   "Carrier_33_Status.10" AT %I2001.2 : Bool;
   "Carrier_33_Status.11" AT %I2001.3 : Bool;
   "Carrier_33_Status.12" AT %I2001.4 : Bool;
   "Carrier_33_Status.13" AT %I2001.5 : Bool;
   "Carrier_33_Status.14" AT %I2001.6 : Bool;
   "Carrier_33_Status.15" AT %I2001.7 : Bool;
   "Carrier_33_SDCFaultCode" AT %IW2002 : Word;   // SDC FAULT CODE
   "Carrier_33_CarrierPosition" AT %ID2004 : DWord;   // CARRIER POSITION
   "Carrier_33_CarrierNumber" AT %IW2008 : Word;   // CARRIER NUMBER
   "Carrier_33_G120DControlWord" AT %IW2010 : Word;   // G120D_STW1_CONTROL
   "Carrier_33_G120DControlWord.0" AT %I2010.0 : Bool;   // Bit_00_ON
   "Carrier_33_G120DControlWord.1" AT %I2010.1 : Bool;   // Bit_01_AUS2_INH
   "Carrier_33_G120DControlWord.2" AT %I2010.2 : Bool;   // Bit_02_AUS3_STOP
   "Carrier_33_G120DControlWord.3" AT %I2010.3 : Bool;   // Bit_03_EN
   "Carrier_33_G120DControlWord.4" AT %I2010.4 : Bool;   // Bit_04_EN_RAMP
   "Carrier_33_G120DControlWord.5" AT %I2010.5 : Bool;   // Bit_05_START_RAMP
   "Carrier_33_G120DControlWord.6" AT %I2010.6 : Bool;   // Bit_06_SETPOINT
   "Carrier_33_G120DControlWord.7" AT %I2010.7 : Bool;   // Bit_07_RESET
   "Carrier_33_G120DControlWord.8" AT %I2011.0 : Bool;   // Bit_08_JOG_R
   "Carrier_33_G120DControlWord.9" AT %I2011.1 : Bool;   // Bit_09_JOG_L
   "Carrier_33_G120DControlWord.10" AT %I2011.2 : Bool;   // Bit_10_CONTR_PLC
   "Carrier_33_G120DControlWord.11" AT %I2011.3 : Bool;   // Bit_11_REVERSE
   "Carrier_33_G120DControlWord.12" AT %I2011.4 : Bool;   // Bit_12_BRAKE_RELEASE
   "Carrier_33_G120DControlWord.13" AT %I2011.5 : Bool;   // Bit_13_DDS
   "Carrier_33_G120DControlWord.14" AT %I2011.6 : Bool;   // Bit_14_DO0
   "Carrier_33_G120DControlWord.15" AT %I2011.7 : Bool;   // Bit_15_DO1
   "Carrier_33_G120DStatusWord" AT %IW2012 : Word;   // G120D_ZSW1_STATUS
   "Carrier_33_G120DStatusWord.0" AT %I2012.0 : Bool;   // Bit_00_READY_RUN
   "Carrier_33_G120DStatusWord.1" AT %I2012.1 : Bool;   // Bit_01_READY_ON
   "Carrier_33_G120DStatusWord.2" AT %I2012.2 : Bool;   // Bit_02_ENABLE
   "Carrier_33_G120DStatusWord.3" AT %I2012.3 : Bool;   // Bit_03_FAULT
   "Carrier_33_G120DStatusWord.4" AT %I2012.4 : Bool;   // Bit_04_OFF2
   "Carrier_33_G120DStatusWord.5" AT %I2012.5 : Bool;   // Bit_05_OFF3
   "Carrier_33_G120DStatusWord.6" AT %I2012.6 : Bool;   // Bit_06_LOCK_OUT
   "Carrier_33_G120DStatusWord.7" AT %I2012.7 : Bool;   // Bit_07_WARN
   "Carrier_33_G120DStatusWord.8" AT %I2013.0 : Bool;   // Bit_08_NO_DEVIATION
   "Carrier_33_G120DStatusWord.9" AT %I2013.1 : Bool;   // Bit_09_CONTR_PLC
   "Carrier_33_G120DStatusWord.10" AT %I2013.2 : Bool;   // Bit_10_F_MAX
   "Carrier_33_G120DStatusWord.11" AT %I2013.3 : Bool;   // Bit_11_LIMIT_REACHED
   "Carrier_33_G120DStatusWord.12" AT %I2013.4 : Bool;   // Bit_12_BRAKE_OPEN
   "Carrier_33_G120DStatusWord.13" AT %I2013.5 : Bool;   // Bit_13_NO_OVERTEMP
   "Carrier_33_G120DStatusWord.14" AT %I2013.6 : Bool;   // Bit_14_CW_CCW
   "Carrier_33_G120DStatusWord.15" AT %I2013.7 : Bool;   // Bit_15_OVERL
   "Carrier_33_Slot2_Input" AT %IW2014 : Word;   // SLOT 2 INPUT WORD
   "Carrier_33_CrashDetectSW" AT %I2014.0 : Bool;   // CRASH DETECT SW
   "Carrier_33_SpareSafetyInput(2_1)" AT %I2014.1 : Bool;   // SPARE SAFETY INPUT
   "Carrier_33_SpareSafetyInput(2_2)" AT %I2014.2 : Bool;   // SPARE SAFETY INPUT
   "Carrier_33_SpareSafetyInput(2_3)" AT %I2014.3 : Bool;   // SPARE SAFETY INPUT
   "Carrier_33_SpareSafetyInput(2_4)" AT %I2014.4 : Bool;   // SPARE SAFETY INPUT
   "Carrier_33_SpareSafetyInput(2_5)" AT %I2014.5 : Bool;   // SPARE SAFETY INPUT
   "Carrier_33_SpareSafetyInput(2_6)" AT %I2014.6 : Bool;   // SPARE SAFETY INPUT
   "Carrier_33_SpareSafetyInput(2_7)" AT %I2014.7 : Bool;   // SPARE SAFETY INPUT
   "Carrier_33_Slot3_SafetyOutput" AT %IW2015 : Word;   // SLOT 3 SAFETY OUTPUT WORD
   "Carrier_33_Crash_Detect_OK" AT %I2015.0 : Bool;   // CARRIER CRASH DETECT
   "Carrier_33_SpareSafetyOutput(3_1)" AT %I2015.1 : Bool;   // SPARE SAFETY OUTPUT
   "Carrier_33_SpareSafetyOutput(3_2)" AT %I2015.2 : Bool;   // SPARE SAFETY OUTPUT
   "Carrier_33_SpareSafetyOutput(3_3)" AT %I2015.3 : Bool;   // SPARE SAFETY OUTPUT
   "Carrier_33_SpareSafetyOutput(3_4)" AT %I2015.4 : Bool;   // SPARE SAFETY OUTPUT
   "Carrier_33_SpareSafetyOutput(3_5)" AT %I2015.5 : Bool;   // SPARE SAFETY OUTPUT
   "Carrier_33_SpareSafetyOutput(3_6)" AT %I2015.6 : Bool;   // SPARE SAFETY OUTPUT
   "Carrier_33_SpareSafetyOutput(3_7)" AT %I2015.7 : Bool;   // SPARE SAFETY OUTPUT
   "Carrier_33_Slot4_Input" AT %IW2016 : Word;   // SLOT 4 INPUT WORD
   "Carrier_33_480VPowerOn_MDCB1" AT %I2016.0 : Bool;   // 480 VAC POWER ON MDCB 1
   "Carrier_33_SpareInput(4_1)" AT %I2016.1 : Bool;   // SPARE INPUT
   "Carrier_33_SpareInput(4_2)" AT %I2016.2 : Bool;   // SPARE INPUT
   "Carrier_33_SitopSelectStatus" AT %I2016.3 : Bool;   // SITOP SELECT STATUS
   "Carrier_33_DCsupplyOnPSCB2" AT %I2016.4 : Bool;   // DC SUPPLY ON PSCB 2
   "Carrier_33_SpareInput(4_5)" AT %I2016.5 : Bool;   // SPARE INPUT
   "Carrier_33_SpareInput(4_6)" AT %I2016.6 : Bool;   // SPARE INPUT
   "Carrier_33_SpareInput(4_7)" AT %I2016.7 : Bool;   // SPARE INPUT
   "Carrier_33_PB1_ProdHoldLH" AT %I2017.0 : Bool;   // PB 1 PRODUCTION HOLD LH
   "Carrier_33_PB2_ResetLH" AT %I2017.1 : Bool;   // PB 2 RESET LH
   "Carrier_33_PB3_ProdHoldRH" AT %I2017.2 : Bool;   // PB 3 PRODUCTION HOLD RH
   "Carrier_33_PB4_ResetRH" AT %I2017.3 : Bool;   // PB 4 RESET RH
   "Carrier_33_SpareInput(4_14)" AT %I2017.4 : Bool;   // SPARE INPUT
   "Carrier_33_SpareInput(4_15)" AT %I2017.5 : Bool;   // SPARE INPUT
   "Carrier_33_SpareInput(4_16)" AT %I2017.6 : Bool;   // SPARE INPUT
   "Carrier_33_SpareInput(4_17)" AT %I2017.7 : Bool;   // SPARE INPUT
   "Carrier_33_Slot5_Output" AT %IW2018 : Word;   // SLOT 5 OUTPUT WORD
   "Carrier_33_IRD400_HMI_24VDC_ENABLE" AT %I2018.0 : Bool;   // IRD 400 PANEL HMI 24V DC POWER
   "Carrier_33_FaultLight_LH" AT %I2018.1 : Bool;   // FAULT LIGHT LH
   "Carrier_33_RunLight_LH" AT %I2018.2 : Bool;   // RUN LIGHT LH
   "Carrier_33_FaultLight_RH" AT %I2018.3 : Bool;   // FAULT LIGHT RH
   "Carrier_33_RunLight_RH" AT %I2018.4 : Bool;   // RUN LIGHT RH
   "Carrier_33_SpareOutput(5_5)" AT %I2018.5 : Bool;   // SPARE OUTPUT
   "Carrier_33_SpareOutput(5_6)" AT %I2018.6 : Bool;   // SPARE OUTPUT
   "Carrier_33_SpareOutput(5_7)" AT %I2018.7 : Bool;   // SPARE OUTPUT
   "Carrier_33_ActualSpeed" AT %IW2020 : Word;   // ACTUAL SPEED
   "Carrier_33_CarrierDriveAlarm" AT %IW2022 : Word;   // CARRIER DRIVE ALARM
   "Carrier_33_CarrierDriveWarning" AT %IW2024 : Word;   // CARRIER DRIVE WARNING
   "Carrier_34_Status" AT %IW2050 : Word;   // CARRIER STATUS WORD
   "Carrier_34_Status.0" AT %I2050.0 : Bool;   // HEARTBEAT
   "Carrier_34_Status.1" AT %I2050.1 : Bool;   // MANUAL
   "Carrier_34_Status.2" AT %I2050.2 : Bool;   // IN_AUTO
   "Carrier_34_Status.3" AT %I2050.3 : Bool;   // POSITIONING_COMPLETE
   "Carrier_34_Status.4" AT %I2050.4 : Bool;   // PRODUCTION HOLD
   "Carrier_34_Status.5" AT %I2050.5 : Bool;   // CARRIER MOVING FORWARD
   "Carrier_34_Status.6" AT %I2050.6 : Bool;   // CARRIER MOVING REVERSE
   "Carrier_34_Status.7" AT %I2050.7 : Bool;   // CARRIER FAULT
   "Carrier_34_Status.8" AT %I2051.0 : Bool;   // CRASH DETECT TRIPPED
   "Carrier_34_Status.9" AT %I2051.1 : Bool;
   "Carrier_34_Status.10" AT %I2051.2 : Bool;
   "Carrier_34_Status.11" AT %I2051.3 : Bool;
   "Carrier_34_Status.12" AT %I2051.4 : Bool;
   "Carrier_34_Status.13" AT %I2051.5 : Bool;
   "Carrier_34_Status.14" AT %I2051.6 : Bool;
   "Carrier_34_Status.15" AT %I2051.7 : Bool;
   "Carrier_34_SDCFaultCode" AT %IW2052 : Word;   // SDC FAULT CODE
   "Carrier_34_CarrierPosition" AT %ID2054 : DWord;   // CARRIER POSITION
   "Carrier_34_CarrierNumber" AT %IW2058 : Word;   // CARRIER NUMBER
   "Carrier_34_G120DControlWord" AT %IW2060 : Word;   // G120D_STW1_CONTROL
   "Carrier_34_G120DControlWord.0" AT %I2060.0 : Bool;   // Bit_00_ON
   "Carrier_34_G120DControlWord.1" AT %I2060.1 : Bool;   // Bit_01_AUS2_INH
   "Carrier_34_G120DControlWord.2" AT %I2060.2 : Bool;   // Bit_02_AUS3_STOP
   "Carrier_34_G120DControlWord.3" AT %I2060.3 : Bool;   // Bit_03_EN
   "Carrier_34_G120DControlWord.4" AT %I2060.4 : Bool;   // Bit_04_EN_RAMP
   "Carrier_34_G120DControlWord.5" AT %I2060.5 : Bool;   // Bit_05_START_RAMP
   "Carrier_34_G120DControlWord.6" AT %I2060.6 : Bool;   // Bit_06_SETPOINT
   "Carrier_34_G120DControlWord.7" AT %I2060.7 : Bool;   // Bit_07_RESET
   "Carrier_34_G120DControlWord.8" AT %I2061.0 : Bool;   // Bit_08_JOG_R
   "Carrier_34_G120DControlWord.9" AT %I2061.1 : Bool;   // Bit_09_JOG_L
   "Carrier_34_G120DControlWord.10" AT %I2061.2 : Bool;   // Bit_10_CONTR_PLC
   "Carrier_34_G120DControlWord.11" AT %I2061.3 : Bool;   // Bit_11_REVERSE
   "Carrier_34_G120DControlWord.12" AT %I2061.4 : Bool;   // Bit_12_BRAKE_RELEASE
   "Carrier_34_G120DControlWord.13" AT %I2061.5 : Bool;   // Bit_13_DDS
   "Carrier_34_G120DControlWord.14" AT %I2061.6 : Bool;   // Bit_14_DO0
   "Carrier_34_G120DControlWord.15" AT %I2061.7 : Bool;   // Bit_15_DO1
   "Carrier_34_G120DStatusWord" AT %IW2062 : Word;   // G120D_ZSW1_STATUS
   "Carrier_34_G120DStatusWord.0" AT %I2062.0 : Bool;   // Bit_00_READY_RUN
   "Carrier_34_G120DStatusWord.1" AT %I2062.1 : Bool;   // Bit_01_READY_ON
   "Carrier_34_G120DStatusWord.2" AT %I2062.2 : Bool;   // Bit_02_ENABLE
   "Carrier_34_G120DStatusWord.3" AT %I2062.3 : Bool;   // Bit_03_FAULT
   "Carrier_34_G120DStatusWord.4" AT %I2062.4 : Bool;   // Bit_04_OFF2
   "Carrier_34_G120DStatusWord.5" AT %I2062.5 : Bool;   // Bit_05_OFF3
   "Carrier_34_G120DStatusWord.6" AT %I2062.6 : Bool;   // Bit_06_LOCK_OUT
   "Carrier_34_G120DStatusWord.7" AT %I2062.7 : Bool;   // Bit_07_WARN
   "Carrier_34_G120DStatusWord.8" AT %I2063.0 : Bool;   // Bit_08_NO_DEVIATION
   "Carrier_34_G120DStatusWord.9" AT %I2063.1 : Bool;   // Bit_09_CONTR_PLC
   "Carrier_34_G120DStatusWord.10" AT %I2063.2 : Bool;   // Bit_10_F_MAX
   "Carrier_34_G120DStatusWord.11" AT %I2063.3 : Bool;   // Bit_11_LIMIT_REACHED
   "Carrier_34_G120DStatusWord.12" AT %I2063.4 : Bool;   // Bit_12_BRAKE_OPEN
   "Carrier_34_G120DStatusWord.13" AT %I2063.5 : Bool;   // Bit_13_NO_OVERTEMP
   "Carrier_34_G120DStatusWord.14" AT %I2063.6 : Bool;   // Bit_14_CW_CCW
   "Carrier_34_G120DStatusWord.15" AT %I2063.7 : Bool;   // Bit_15_OVERL
   "Carrier_34_Slot2_Input" AT %IW2064 : Word;   // SLOT 2 INPUT WORD
   "Carrier_34_CrashDetectSW" AT %I2064.0 : Bool;   // CRASH DETECT SW
   "Carrier_34_SpareSafetyInput(2_1)" AT %I2064.1 : Bool;   // SPARE SAFETY INPUT
   "Carrier_34_SpareSafetyInput(2_2)" AT %I2064.2 : Bool;   // SPARE SAFETY INPUT
   "Carrier_34_SpareSafetyInput(2_3)" AT %I2064.3 : Bool;   // SPARE SAFETY INPUT
   "Carrier_34_SpareSafetyInput(2_4)" AT %I2064.4 : Bool;   // SPARE SAFETY INPUT
   "Carrier_34_SpareSafetyInput(2_5)" AT %I2064.5 : Bool;   // SPARE SAFETY INPUT
   "Carrier_34_SpareSafetyInput(2_6)" AT %I2064.6 : Bool;   // SPARE SAFETY INPUT
   "Carrier_34_SpareSafetyInput(2_7)" AT %I2064.7 : Bool;   // SPARE SAFETY INPUT
   "Carrier_34_Slot3_SafetyOutput" AT %IW2065 : Word;   // SLOT 3 SAFETY OUTPUT WORD
   "Carrier_34_Crash_Detect_OK" AT %I2065.0 : Bool;   // CARRIER CRASH DETECT
   "Carrier_34_SpareSafetyOutput(3_1)" AT %I2065.1 : Bool;   // SPARE SAFETY OUTPUT
   "Carrier_34_SpareSafetyOutput(3_2)" AT %I2065.2 : Bool;   // SPARE SAFETY OUTPUT
   "Carrier_34_SpareSafetyOutput(3_3)" AT %I2065.3 : Bool;   // SPARE SAFETY OUTPUT
   "Carrier_34_SpareSafetyOutput(3_4)" AT %I2065.4 : Bool;   // SPARE SAFETY OUTPUT
   "Carrier_34_SpareSafetyOutput(3_5)" AT %I2065.5 : Bool;   // SPARE SAFETY OUTPUT
   "Carrier_34_SpareSafetyOutput(3_6)" AT %I2065.6 : Bool;   // SPARE SAFETY OUTPUT
   "Carrier_34_SpareSafetyOutput(3_7)" AT %I2065.7 : Bool;   // SPARE SAFETY OUTPUT
   "Carrier_34_Slot4_Input" AT %IW2066 : Word;   // SLOT 4 INPUT WORD
   "Carrier_34_480VPowerOn_MDCB1" AT %I2066.0 : Bool;   // 480 VAC POWER ON MDCB 1
   "Carrier_34_SpareInput(4_1)" AT %I2066.1 : Bool;   // SPARE INPUT
   "Carrier_34_SpareInput(4_2)" AT %I2066.2 : Bool;   // SPARE INPUT
   "Carrier_34_SitopSelectStatus" AT %I2066.3 : Bool;   // SITOP SELECT STATUS
   "Carrier_34_DCsupplyOnPSCB2" AT %I2066.4 : Bool;   // DC SUPPLY ON PSCB 2
   "Carrier_34_SpareInput(4_5)" AT %I2066.5 : Bool;   // SPARE INPUT
   "Carrier_34_SpareInput(4_6)" AT %I2066.6 : Bool;   // SPARE INPUT
   "Carrier_34_SpareInput(4_7)" AT %I2066.7 : Bool;   // SPARE INPUT
   "Carrier_34_PB1_ProdHoldLH" AT %I2067.0 : Bool;   // PB 1 PRODUCTION HOLD LH
   "Carrier_34_PB2_ResetLH" AT %I2067.1 : Bool;   // PB 2 RESET LH
   "Carrier_34_PB3_ProdHoldRH" AT %I2067.2 : Bool;   // PB 3 PRODUCTION HOLD RH
   "Carrier_34_PB4_ResetRH" AT %I2067.3 : Bool;   // PB 4 RESET RH
   "Carrier_34_SpareInput(4_14)" AT %I2067.4 : Bool;   // SPARE INPUT
   "Carrier_34_SpareInput(4_15)" AT %I2067.5 : Bool;   // SPARE INPUT
   "Carrier_34_SpareInput(4_16)" AT %I2067.6 : Bool;   // SPARE INPUT
   "Carrier_34_SpareInput(4_17)" AT %I2067.7 : Bool;   // SPARE INPUT
   "Carrier_34_Slot5_Output" AT %IW2068 : Word;   // SLOT 5 OUTPUT WORD
   "Carrier_34_IRD400_HMI_24VDC_ENABLE" AT %I2068.0 : Bool;   // IRD 400 PANEL HMI 24V DC POWER
   "Carrier_34_FaultLight_LH" AT %I2068.1 : Bool;   // FAULT LIGHT LH
   "Carrier_34_RunLight_LH" AT %I2068.2 : Bool;   // RUN LIGHT LH
   "Carrier_34_FaultLight_RH" AT %I2068.3 : Bool;   // FAULT LIGHT RH
   "Carrier_34_RunLight_RH" AT %I2068.4 : Bool;   // RUN LIGHT RH
   "Carrier_34_SpareOutput(5_5)" AT %I2068.5 : Bool;   // SPARE OUTPUT
   "Carrier_34_SpareOutput(5_6)" AT %I2068.6 : Bool;   // SPARE OUTPUT
   "Carrier_34_SpareOutput(5_7)" AT %I2068.7 : Bool;   // SPARE OUTPUT
   "Carrier_34_ActualSpeed" AT %IW2070 : Word;   // ACTUAL SPEED
   "Carrier_34_CarrierDriveAlarm" AT %IW2072 : Word;   // CARRIER DRIVE ALARM
   "Carrier_34_CarrierDriveWarning" AT %IW2074 : Word;   // CARRIER DRIVE WARNING
   "Carrier_35_Status" AT %IW2100 : Word;   // CARRIER STATUS WORD
   "Carrier_35_Status.0" AT %I2100.0 : Bool;   // HEARTBEAT
   "Carrier_35_Status.1" AT %I2100.1 : Bool;   // MANUAL
   "Carrier_35_Status.2" AT %I2100.2 : Bool;   // IN_AUTO
   "Carrier_35_Status.3" AT %I2100.3 : Bool;   // POSITIONING_COMPLETE
   "Carrier_35_Status.4" AT %I2100.4 : Bool;   // PRODUCTION HOLD
   "Carrier_35_Status.5" AT %I2100.5 : Bool;   // CARRIER MOVING FORWARD
   "Carrier_35_Status.6" AT %I2100.6 : Bool;   // CARRIER MOVING REVERSE
   "Carrier_35_Status.7" AT %I2100.7 : Bool;   // CARRIER FAULT
   "Carrier_35_Status.8" AT %I2101.0 : Bool;   // CRASH DETECT TRIPPED
   "Carrier_35_Status.9" AT %I2101.1 : Bool;
   "Carrier_35_Status.10" AT %I2101.2 : Bool;
   "Carrier_35_Status.11" AT %I2101.3 : Bool;
   "Carrier_35_Status.12" AT %I2101.4 : Bool;
   "Carrier_35_Status.13" AT %I2101.5 : Bool;
   "Carrier_35_Status.14" AT %I2101.6 : Bool;
   "Carrier_35_Status.15" AT %I2101.7 : Bool;
   "Carrier_35_SDCFaultCode" AT %IW2102 : Word;   // SDC FAULT CODE
   "Carrier_35_CarrierPosition" AT %ID2104 : DWord;   // CARRIER POSITION
   "Carrier_35_CarrierNumber" AT %IW2108 : Word;   // CARRIER NUMBER
   "Carrier_35_G120DControlWord" AT %IW2110 : Word;   // G120D_STW1_CONTROL
   "Carrier_35_G120DControlWord.0" AT %I2110.0 : Bool;   // Bit_00_ON
   "Carrier_35_G120DControlWord.1" AT %I2110.1 : Bool;   // Bit_01_AUS2_INH
   "Carrier_35_G120DControlWord.2" AT %I2110.2 : Bool;   // Bit_02_AUS3_STOP
   "Carrier_35_G120DControlWord.3" AT %I2110.3 : Bool;   // Bit_03_EN
   "Carrier_35_G120DControlWord.4" AT %I2110.4 : Bool;   // Bit_04_EN_RAMP
   "Carrier_35_G120DControlWord.5" AT %I2110.5 : Bool;   // Bit_05_START_RAMP
   "Carrier_35_G120DControlWord.6" AT %I2110.6 : Bool;   // Bit_06_SETPOINT
   "Carrier_35_G120DControlWord.7" AT %I2110.7 : Bool;   // Bit_07_RESET
   "Carrier_35_G120DControlWord.8" AT %I2111.0 : Bool;   // Bit_08_JOG_R
   "Carrier_35_G120DControlWord.9" AT %I2111.1 : Bool;   // Bit_09_JOG_L
   "Carrier_35_G120DControlWord.10" AT %I2111.2 : Bool;   // Bit_10_CONTR_PLC
   "Carrier_35_G120DControlWord.11" AT %I2111.3 : Bool;   // Bit_11_REVERSE
   "Carrier_35_G120DControlWord.12" AT %I2111.4 : Bool;   // Bit_12_BRAKE_RELEASE
   "Carrier_35_G120DControlWord.13" AT %I2111.5 : Bool;   // Bit_13_DDS
   "Carrier_35_G120DControlWord.14" AT %I2111.6 : Bool;   // Bit_14_DO0
   "Carrier_35_G120DControlWord.15" AT %I2111.7 : Bool;   // Bit_15_DO1
   "Carrier_35_G120DStatusWord" AT %IW2112 : Word;   // G120D_ZSW1_STATUS
   "Carrier_35_G120DStatusWord.0" AT %I2112.0 : Bool;   // Bit_00_READY_RUN
   "Carrier_35_G120DStatusWord.1" AT %I2112.1 : Bool;   // Bit_01_READY_ON
   "Carrier_35_G120DStatusWord.2" AT %I2112.2 : Bool;   // Bit_02_ENABLE
   "Carrier_35_G120DStatusWord.3" AT %I2112.3 : Bool;   // Bit_03_FAULT
   "Carrier_35_G120DStatusWord.4" AT %I2112.4 : Bool;   // Bit_04_OFF2
   "Carrier_35_G120DStatusWord.5" AT %I2112.5 : Bool;   // Bit_05_OFF3
   "Carrier_35_G120DStatusWord.6" AT %I2112.6 : Bool;   // Bit_06_LOCK_OUT
   "Carrier_35_G120DStatusWord.7" AT %I2112.7 : Bool;   // Bit_07_WARN
   "Carrier_35_G120DStatusWord.8" AT %I2113.0 : Bool;   // Bit_08_NO_DEVIATION
   "Carrier_35_G120DStatusWord.9" AT %I2113.1 : Bool;   // Bit_09_CONTR_PLC
   "Carrier_35_G120DStatusWord.10" AT %I2113.2 : Bool;   // Bit_10_F_MAX
   "Carrier_35_G120DStatusWord.11" AT %I2113.3 : Bool;   // Bit_11_LIMIT_REACHED
   "Carrier_35_G120DStatusWord.12" AT %I2113.4 : Bool;   // Bit_12_BRAKE_OPEN
   "Carrier_35_G120DStatusWord.13" AT %I2113.5 : Bool;   // Bit_13_NO_OVERTEMP
   "Carrier_35_G120DStatusWord.14" AT %I2113.6 : Bool;   // Bit_14_CW_CCW
   "Carrier_35_G120DStatusWord.15" AT %I2113.7 : Bool;   // Bit_15_OVERL
   "Carrier_35_Slot2_Input" AT %IW2114 : Word;   // SLOT 2 INPUT WORD
   "Carrier_35_CrashDetectSW" AT %I2114.0 : Bool;   // CRASH DETECT SW
   "Carrier_35_SpareSafetyInput(2_1)" AT %I2114.1 : Bool;   // SPARE SAFETY INPUT
   "Carrier_35_SpareSafetyInput(2_2)" AT %I2114.2 : Bool;   // SPARE SAFETY INPUT
   "Carrier_35_SpareSafetyInput(2_3)" AT %I2114.3 : Bool;   // SPARE SAFETY INPUT
   "Carrier_35_SpareSafetyInput(2_4)" AT %I2114.4 : Bool;   // SPARE SAFETY INPUT
   "Carrier_35_SpareSafetyInput(2_5)" AT %I2114.5 : Bool;   // SPARE SAFETY INPUT
   "Carrier_35_SpareSafetyInput(2_6)" AT %I2114.6 : Bool;   // SPARE SAFETY INPUT
   "Carrier_35_SpareSafetyInput(2_7)" AT %I2114.7 : Bool;   // SPARE SAFETY INPUT
   "Carrier_35_Slot3_SafetyOutput" AT %IW2115 : Word;   // SLOT 3 SAFETY OUTPUT WORD
   "Carrier_35_Crash_Detect_OK" AT %I2115.0 : Bool;   // CARRIER CRASH DETECT
   "Carrier_35_SpareSafetyOutput(3_1)" AT %I2115.1 : Bool;   // SPARE SAFETY OUTPUT
   "Carrier_35_SpareSafetyOutput(3_2)" AT %I2115.2 : Bool;   // SPARE SAFETY OUTPUT
   "Carrier_35_SpareSafetyOutput(3_3)" AT %I2115.3 : Bool;   // SPARE SAFETY OUTPUT
   "Carrier_35_SpareSafetyOutput(3_4)" AT %I2115.4 : Bool;   // SPARE SAFETY OUTPUT
   "Carrier_35_SpareSafetyOutput(3_5)" AT %I2115.5 : Bool;   // SPARE SAFETY OUTPUT
   "Carrier_35_SpareSafetyOutput(3_6)" AT %I2115.6 : Bool;   // SPARE SAFETY OUTPUT
   "Carrier_35_SpareSafetyOutput(3_7)" AT %I2115.7 : Bool;   // SPARE SAFETY OUTPUT
   "Carrier_35_Slot4_Input" AT %IW2116 : Word;   // SLOT 4 INPUT WORD
   "Carrier_35_480VPowerOn_MDCB1" AT %I2116.0 : Bool;   // 480 VAC POWER ON MDCB 1
   "Carrier_35_SpareInput(4_1)" AT %I2116.1 : Bool;   // SPARE INPUT
   "Carrier_35_SpareInput(4_2)" AT %I2116.2 : Bool;   // SPARE INPUT
   "Carrier_35_SitopSelectStatus" AT %I2116.3 : Bool;   // SITOP SELECT STATUS
   "Carrier_35_DCsupplyOnPSCB2" AT %I2116.4 : Bool;   // DC SUPPLY ON PSCB 2
   "Carrier_35_SpareInput(4_5)" AT %I2116.5 : Bool;   // SPARE INPUT
   "Carrier_35_SpareInput(4_6)" AT %I2116.6 : Bool;   // SPARE INPUT
   "Carrier_35_SpareInput(4_7)" AT %I2116.7 : Bool;   // SPARE INPUT
   "Carrier_35_PB1_ProdHoldLH" AT %I2117.0 : Bool;   // PB 1 PRODUCTION HOLD LH
   "Carrier_35_PB2_ResetLH" AT %I2117.1 : Bool;   // PB 2 RESET LH
   "Carrier_35_PB3_ProdHoldRH" AT %I2117.2 : Bool;   // PB 3 PRODUCTION HOLD RH
   "Carrier_35_PB4_ResetRH" AT %I2117.3 : Bool;   // PB 4 RESET RH
   "Carrier_35_SpareInput(4_14)" AT %I2117.4 : Bool;   // SPARE INPUT
   "Carrier_35_SpareInput(4_15)" AT %I2117.5 : Bool;   // SPARE INPUT
   "Carrier_35_SpareInput(4_16)" AT %I2117.6 : Bool;   // SPARE INPUT
   "Carrier_35_SpareInput(4_17)" AT %I2117.7 : Bool;   // SPARE INPUT
   "Carrier_35_Slot5_Output" AT %IW2118 : Word;   // SLOT 5 OUTPUT WORD
   "Carrier_35_IRD400_HMI_24VDC_ENABLE" AT %I2118.0 : Bool;   // IRD 400 PANEL HMI 24V DC POWER
   "Carrier_35_FaultLight_LH" AT %I2118.1 : Bool;   // FAULT LIGHT LH
   "Carrier_35_RunLight_LH" AT %I2118.2 : Bool;   // RUN LIGHT LH
   "Carrier_35_FaultLight_RH" AT %I2118.3 : Bool;   // FAULT LIGHT RH
   "Carrier_35_RunLight_RH" AT %I2118.4 : Bool;   // RUN LIGHT RH
   "Carrier_35_SpareOutput(5_5)" AT %I2118.5 : Bool;   // SPARE OUTPUT
   "Carrier_35_SpareOutput(5_6)" AT %I2118.6 : Bool;   // SPARE OUTPUT
   "Carrier_35_SpareOutput(5_7)" AT %I2118.7 : Bool;   // SPARE OUTPUT
   "Carrier_35_ActualSpeed" AT %IW2120 : Word;   // ACTUAL SPEED
   "Carrier_35_CarrierDriveAlarm" AT %IW2122 : Word;   // CARRIER DRIVE ALARM
   "Carrier_35_CarrierDriveWarning" AT %IW2124 : Word;   // CARRIER DRIVE WARNING
   "Carrier_36_Status" AT %IW2150 : Word;   // CARRIER STATUS WORD
   "Carrier_36_Status.0" AT %I2150.0 : Bool;   // HEARTBEAT
   "Carrier_36_Status.1" AT %I2150.1 : Bool;   // MANUAL
   "Carrier_36_Status.2" AT %I2150.2 : Bool;   // IN_AUTO
   "Carrier_36_Status.3" AT %I2150.3 : Bool;   // POSITIONING_COMPLETE
   "Carrier_36_Status.4" AT %I2150.4 : Bool;   // PRODUCTION HOLD
   "Carrier_36_Status.5" AT %I2150.5 : Bool;   // CARRIER MOVING FORWARD
   "Carrier_36_Status.6" AT %I2150.6 : Bool;   // CARRIER MOVING REVERSE
   "Carrier_36_Status.7" AT %I2150.7 : Bool;   // CARRIER FAULT
   "Carrier_36_Status.8" AT %I2151.0 : Bool;   // CRASH DETECT TRIPPED
   "Carrier_36_Status.9" AT %I2151.1 : Bool;
   "Carrier_36_Status.10" AT %I2151.2 : Bool;
   "Carrier_36_Status.11" AT %I2151.3 : Bool;
   "Carrier_36_Status.12" AT %I2151.4 : Bool;
   "Carrier_36_Status.13" AT %I2151.5 : Bool;
   "Carrier_36_Status.14" AT %I2151.6 : Bool;
   "Carrier_36_Status.15" AT %I2151.7 : Bool;
   "Carrier_36_SDCFaultCode" AT %IW2152 : Word;   // SDC FAULT CODE
   "Carrier_36_CarrierPosition" AT %ID2154 : DWord;   // CARRIER POSITION
   "Carrier_36_CarrierNumber" AT %IW2158 : Word;   // CARRIER NUMBER
   "Carrier_36_G120DControlWord" AT %IW2160 : Word;   // G120D_STW1_CONTROL
   "Carrier_36_G120DControlWord.0" AT %I2160.0 : Bool;   // Bit_00_ON
   "Carrier_36_G120DControlWord.1" AT %I2160.1 : Bool;   // Bit_01_AUS2_INH
   "Carrier_36_G120DControlWord.2" AT %I2160.2 : Bool;   // Bit_02_AUS3_STOP
   "Carrier_36_G120DControlWord.3" AT %I2160.3 : Bool;   // Bit_03_EN
   "Carrier_36_G120DControlWord.4" AT %I2160.4 : Bool;   // Bit_04_EN_RAMP
   "Carrier_36_G120DControlWord.5" AT %I2160.5 : Bool;   // Bit_05_START_RAMP
   "Carrier_36_G120DControlWord.6" AT %I2160.6 : Bool;   // Bit_06_SETPOINT
   "Carrier_36_G120DControlWord.7" AT %I2160.7 : Bool;   // Bit_07_RESET
   "Carrier_36_G120DControlWord.8" AT %I2161.0 : Bool;   // Bit_08_JOG_R
   "Carrier_36_G120DControlWord.9" AT %I2161.1 : Bool;   // Bit_09_JOG_L
   "Carrier_36_G120DControlWord.10" AT %I2161.2 : Bool;   // Bit_10_CONTR_PLC
   "Carrier_36_G120DControlWord.11" AT %I2161.3 : Bool;   // Bit_11_REVERSE
   "Carrier_36_G120DControlWord.12" AT %I2161.4 : Bool;   // Bit_12_BRAKE_RELEASE
   "Carrier_36_G120DControlWord.13" AT %I2161.5 : Bool;   // Bit_13_DDS
   "Carrier_36_G120DControlWord.14" AT %I2161.6 : Bool;   // Bit_14_DO0
   "Carrier_36_G120DControlWord.15" AT %I2161.7 : Bool;   // Bit_15_DO1
   "Carrier_36_G120DStatusWord" AT %IW2162 : Word;   // G120D_ZSW1_STATUS
   "Carrier_36_G120DStatusWord.0" AT %I2162.0 : Bool;   // Bit_00_READY_RUN
   "Carrier_36_G120DStatusWord.1" AT %I2162.1 : Bool;   // Bit_01_READY_ON
   "Carrier_36_G120DStatusWord.2" AT %I2162.2 : Bool;   // Bit_02_ENABLE
   "Carrier_36_G120DStatusWord.3" AT %I2162.3 : Bool;   // Bit_03_FAULT
   "Carrier_36_G120DStatusWord.4" AT %I2162.4 : Bool;   // Bit_04_OFF2
   "Carrier_36_G120DStatusWord.5" AT %I2162.5 : Bool;   // Bit_05_OFF3
   "Carrier_36_G120DStatusWord.6" AT %I2162.6 : Bool;   // Bit_06_LOCK_OUT
   "Carrier_36_G120DStatusWord.7" AT %I2162.7 : Bool;   // Bit_07_WARN
   "Carrier_36_G120DStatusWord.8" AT %I2163.0 : Bool;   // Bit_08_NO_DEVIATION
   "Carrier_36_G120DStatusWord.9" AT %I2163.1 : Bool;   // Bit_09_CONTR_PLC
   "Carrier_36_G120DStatusWord.10" AT %I2163.2 : Bool;   // Bit_10_F_MAX
   "Carrier_36_G120DStatusWord.11" AT %I2163.3 : Bool;   // Bit_11_LIMIT_REACHED
   "Carrier_36_G120DStatusWord.12" AT %I2163.4 : Bool;   // Bit_12_BRAKE_OPEN
   "Carrier_36_G120DStatusWord.13" AT %I2163.5 : Bool;   // Bit_13_NO_OVERTEMP
   "Carrier_36_G120DStatusWord.14" AT %I2163.6 : Bool;   // Bit_14_CW_CCW
   "Carrier_36_G120DStatusWord.15" AT %I2163.7 : Bool;   // Bit_15_OVERL
   "Carrier_36_Slot2_Input" AT %IW2164 : Word;   // SLOT 2 INPUT WORD
   "Carrier_36_CrashDetectSW" AT %I2164.0 : Bool;   // CRASH DETECT SW
   "Carrier_36_SpareSafetyInput(2_1)" AT %I2164.1 : Bool;   // SPARE SAFETY INPUT
   "Carrier_36_SpareSafetyInput(2_2)" AT %I2164.2 : Bool;   // SPARE SAFETY INPUT
   "Carrier_36_SpareSafetyInput(2_3)" AT %I2164.3 : Bool;   // SPARE SAFETY INPUT
   "Carrier_36_SpareSafetyInput(2_4)" AT %I2164.4 : Bool;   // SPARE SAFETY INPUT
   "Carrier_36_SpareSafetyInput(2_5)" AT %I2164.5 : Bool;   // SPARE SAFETY INPUT
   "Carrier_36_SpareSafetyInput(2_6)" AT %I2164.6 : Bool;   // SPARE SAFETY INPUT
   "Carrier_36_SpareSafetyInput(2_7)" AT %I2164.7 : Bool;   // SPARE SAFETY INPUT
   "Carrier_36_Slot3_SafetyOutput" AT %IW2165 : Word;   // SLOT 3 SAFETY OUTPUT WORD
   "Carrier_36_Crash_Detect_OK" AT %I2165.0 : Bool;   // CARRIER CRASH DETECT
   "Carrier_36_SpareSafetyOutput(3_1)" AT %I2165.1 : Bool;   // SPARE SAFETY OUTPUT
   "Carrier_36_SpareSafetyOutput(3_2)" AT %I2165.2 : Bool;   // SPARE SAFETY OUTPUT
   "Carrier_36_SpareSafetyOutput(3_3)" AT %I2165.3 : Bool;   // SPARE SAFETY OUTPUT
   "Carrier_36_SpareSafetyOutput(3_4)" AT %I2165.4 : Bool;   // SPARE SAFETY OUTPUT
   "Carrier_36_SpareSafetyOutput(3_5)" AT %I2165.5 : Bool;   // SPARE SAFETY OUTPUT
   "Carrier_36_SpareSafetyOutput(3_6)" AT %I2165.6 : Bool;   // SPARE SAFETY OUTPUT
   "Carrier_36_SpareSafetyOutput(3_7)" AT %I2165.7 : Bool;   // SPARE SAFETY OUTPUT
   "Carrier_36_Slot4_Input" AT %IW2166 : Word;   // SLOT 4 INPUT WORD
   "Carrier_36_480VPowerOn_MDCB1" AT %I2166.0 : Bool;   // 480 VAC POWER ON MDCB 1
   "Carrier_36_SpareInput(4_1)" AT %I2166.1 : Bool;   // SPARE INPUT
   "Carrier_36_SpareInput(4_2)" AT %I2166.2 : Bool;   // SPARE INPUT
   "Carrier_36_SitopSelectStatus" AT %I2166.3 : Bool;   // SITOP SELECT STATUS
   "Carrier_36_DCsupplyOnPSCB2" AT %I2166.4 : Bool;   // DC SUPPLY ON PSCB 2
   "Carrier_36_SpareInput(4_5)" AT %I2166.5 : Bool;   // SPARE INPUT
   "Carrier_36_SpareInput(4_6)" AT %I2166.6 : Bool;   // SPARE INPUT
   "Carrier_36_SpareInput(4_7)" AT %I2166.7 : Bool;   // SPARE INPUT
   "Carrier_36_PB1_ProdHoldLH" AT %I2167.0 : Bool;   // PB 1 PRODUCTION HOLD LH
   "Carrier_36_PB2_ResetLH" AT %I2167.1 : Bool;   // PB 2 RESET LH
   "Carrier_36_PB3_ProdHoldRH" AT %I2167.2 : Bool;   // PB 3 PRODUCTION HOLD RH
   "Carrier_36_PB4_ResetRH" AT %I2167.3 : Bool;   // PB 4 RESET RH
   "Carrier_36_SpareInput(4_14)" AT %I2167.4 : Bool;   // SPARE INPUT
   "Carrier_36_SpareInput(4_15)" AT %I2167.5 : Bool;   // SPARE INPUT
   "Carrier_36_SpareInput(4_16)" AT %I2167.6 : Bool;   // SPARE INPUT
   "Carrier_36_SpareInput(4_17)" AT %I2167.7 : Bool;   // SPARE INPUT
   "Carrier_36_Slot5_Output" AT %IW2168 : Word;   // SLOT 5 OUTPUT WORD
   "Carrier_36_IRD400_HMI_24VDC_ENABLE" AT %I2168.0 : Bool;   // IRD 400 PANEL HMI 24V DC POWER
   "Carrier_36_FaultLight_LH" AT %I2168.1 : Bool;   // FAULT LIGHT LH
   "Carrier_36_RunLight_LH" AT %I2168.2 : Bool;   // RUN LIGHT LH
   "Carrier_36_FaultLight_RH" AT %I2168.3 : Bool;   // FAULT LIGHT RH
   "Carrier_36_RunLight_RH" AT %I2168.4 : Bool;   // RUN LIGHT RH
   "Carrier_36_SpareOutput(5_5)" AT %I2168.5 : Bool;   // SPARE OUTPUT
   "Carrier_36_SpareOutput(5_6)" AT %I2168.6 : Bool;   // SPARE OUTPUT
   "Carrier_36_SpareOutput(5_7)" AT %I2168.7 : Bool;   // SPARE OUTPUT
   "Carrier_36_ActualSpeed" AT %IW2170 : Word;   // ACTUAL SPEED
   "Carrier_36_CarrierDriveAlarm" AT %IW2172 : Word;   // CARRIER DRIVE ALARM
   "Carrier_36_CarrierDriveWarning" AT %IW2174 : Word;   // CARRIER DRIVE WARNING
   "Carrier_37_Status" AT %IW2200 : Word;   // CARRIER STATUS WORD
   "Carrier_37_Status.0" AT %I2200.0 : Bool;   // HEARTBEAT
   "Carrier_37_Status.1" AT %I2200.1 : Bool;   // MANUAL
   "Carrier_37_Status.2" AT %I2200.2 : Bool;   // IN_AUTO
   "Carrier_37_Status.3" AT %I2200.3 : Bool;   // POSITIONING_COMPLETE
   "Carrier_37_Status.4" AT %I2200.4 : Bool;   // PRODUCTION HOLD
   "Carrier_37_Status.5" AT %I2200.5 : Bool;   // CARRIER MOVING FORWARD
   "Carrier_37_Status.6" AT %I2200.6 : Bool;   // CARRIER MOVING REVERSE
   "Carrier_37_Status.7" AT %I2200.7 : Bool;   // CARRIER FAULT
   "Carrier_37_Status.8" AT %I2201.0 : Bool;   // CRASH DETECT TRIPPED
   "Carrier_37_Status.9" AT %I2201.1 : Bool;
   "Carrier_37_Status.10" AT %I2201.2 : Bool;
   "Carrier_37_Status.11" AT %I2201.3 : Bool;
   "Carrier_37_Status.12" AT %I2201.4 : Bool;
   "Carrier_37_Status.13" AT %I2201.5 : Bool;
   "Carrier_37_Status.14" AT %I2201.6 : Bool;
   "Carrier_37_Status.15" AT %I2201.7 : Bool;
   "Carrier_37_SDCFaultCode" AT %IW2202 : Word;   // SDC FAULT CODE
   "Carrier_37_CarrierPosition" AT %ID2204 : DWord;   // CARRIER POSITION
   "Carrier_37_CarrierNumber" AT %IW2208 : Word;   // CARRIER NUMBER
   "Carrier_37_G120DControlWord" AT %IW2210 : Word;   // G120D_STW1_CONTROL
   "Carrier_37_G120DControlWord.0" AT %I2210.0 : Bool;   // Bit_00_ON
   "Carrier_37_G120DControlWord.1" AT %I2210.1 : Bool;   // Bit_01_AUS2_INH
   "Carrier_37_G120DControlWord.2" AT %I2210.2 : Bool;   // Bit_02_AUS3_STOP
   "Carrier_37_G120DControlWord.3" AT %I2210.3 : Bool;   // Bit_03_EN
   "Carrier_37_G120DControlWord.4" AT %I2210.4 : Bool;   // Bit_04_EN_RAMP
   "Carrier_37_G120DControlWord.5" AT %I2210.5 : Bool;   // Bit_05_START_RAMP
   "Carrier_37_G120DControlWord.6" AT %I2210.6 : Bool;   // Bit_06_SETPOINT
   "Carrier_37_G120DControlWord.7" AT %I2210.7 : Bool;   // Bit_07_RESET
   "Carrier_37_G120DControlWord.8" AT %I2211.0 : Bool;   // Bit_08_JOG_R
   "Carrier_37_G120DControlWord.9" AT %I2211.1 : Bool;   // Bit_09_JOG_L
   "Carrier_37_G120DControlWord.10" AT %I2211.2 : Bool;   // Bit_10_CONTR_PLC
   "Carrier_37_G120DControlWord.11" AT %I2211.3 : Bool;   // Bit_11_REVERSE
   "Carrier_37_G120DControlWord.12" AT %I2211.4 : Bool;   // Bit_12_BRAKE_RELEASE
   "Carrier_37_G120DControlWord.13" AT %I2211.5 : Bool;   // Bit_13_DDS
   "Carrier_37_G120DControlWord.14" AT %I2211.6 : Bool;   // Bit_14_DO0
   "Carrier_37_G120DControlWord.15" AT %I2211.7 : Bool;   // Bit_15_DO1
   "Carrier_37_G120DStatusWord" AT %IW2212 : Word;   // G120D_ZSW1_STATUS
   "Carrier_37_G120DStatusWord.0" AT %I2212.0 : Bool;   // Bit_00_READY_RUN
   "Carrier_37_G120DStatusWord.1" AT %I2212.1 : Bool;   // Bit_01_READY_ON
   "Carrier_37_G120DStatusWord.2" AT %I2212.2 : Bool;   // Bit_02_ENABLE
   "Carrier_37_G120DStatusWord.3" AT %I2212.3 : Bool;   // Bit_03_FAULT
   "Carrier_37_G120DStatusWord.4" AT %I2212.4 : Bool;   // Bit_04_OFF2
   "Carrier_37_G120DStatusWord.5" AT %I2212.5 : Bool;   // Bit_05_OFF3
   "Carrier_37_G120DStatusWord.6" AT %I2212.6 : Bool;   // Bit_06_LOCK_OUT
   "Carrier_37_G120DStatusWord.7" AT %I2212.7 : Bool;   // Bit_07_WARN
   "Carrier_37_G120DStatusWord.8" AT %I2213.0 : Bool;   // Bit_08_NO_DEVIATION
   "Carrier_37_G120DStatusWord.9" AT %I2213.1 : Bool;   // Bit_09_CONTR_PLC
   "Carrier_37_G120DStatusWord.10" AT %I2213.2 : Bool;   // Bit_10_F_MAX
   "Carrier_37_G120DStatusWord.11" AT %I2213.3 : Bool;   // Bit_11_LIMIT_REACHED
   "Carrier_37_G120DStatusWord.12" AT %I2213.4 : Bool;   // Bit_12_BRAKE_OPEN
   "Carrier_37_G120DStatusWord.13" AT %I2213.5 : Bool;   // Bit_13_NO_OVERTEMP
   "Carrier_37_G120DStatusWord.14" AT %I2213.6 : Bool;   // Bit_14_CW_CCW
   "Carrier_37_G120DStatusWord.15" AT %I2213.7 : Bool;   // Bit_15_OVERL
   "Carrier_37_Slot2_Input" AT %IW2214 : Word;   // SLOT 2 INPUT WORD
   "Carrier_37_CrashDetectSW" AT %I2214.0 : Bool;   // CRASH DETECT SW
   "Carrier_37_SpareSafetyInput(2_1)" AT %I2214.1 : Bool;   // SPARE SAFETY INPUT
   "Carrier_37_SpareSafetyInput(2_2)" AT %I2214.2 : Bool;   // SPARE SAFETY INPUT
   "Carrier_37_SpareSafetyInput(2_3)" AT %I2214.3 : Bool;   // SPARE SAFETY INPUT
   "Carrier_37_SpareSafetyInput(2_4)" AT %I2214.4 : Bool;   // SPARE SAFETY INPUT
   "Carrier_37_SpareSafetyInput(2_5)" AT %I2214.5 : Bool;   // SPARE SAFETY INPUT
   "Carrier_37_SpareSafetyInput(2_6)" AT %I2214.6 : Bool;   // SPARE SAFETY INPUT
   "Carrier_37_SpareSafetyInput(2_7)" AT %I2214.7 : Bool;   // SPARE SAFETY INPUT
   "Carrier_37_Slot3_SafetyOutput" AT %IW2215 : Word;   // SLOT 3 SAFETY OUTPUT WORD
   "Carrier_37_Crash_Detect_OK" AT %I2215.0 : Bool;   // CARRIER CRASH DETECT
   "Carrier_37_SpareSafetyOutput(3_1)" AT %I2215.1 : Bool;   // SPARE SAFETY OUTPUT
   "Carrier_37_SpareSafetyOutput(3_2)" AT %I2215.2 : Bool;   // SPARE SAFETY OUTPUT
   "Carrier_37_SpareSafetyOutput(3_3)" AT %I2215.3 : Bool;   // SPARE SAFETY OUTPUT